   1118: 'Carrier 17 Power unit: Phase failure motor cable', class No Acknowledgement, trigger "DB302_HMI_Faults_Carrier17_Faults_1" bit 13
   1119: 'Carrier 17 Power unit: Ground fault', class No Acknowledgement, trigger "DB302_HMI_Faults_Carrier17_Faults_1" bit 14
   1120: 'Spare_Fault_1120', class No Acknowledgement, trigger "DB302_HMI_Faults_Carrier17_Faults_1" bit 15
   1121: 'Carrier 17 Motion Off Fault', class No Acknowledgement, trigger "DB302_HMI_Faults_Carrier17_Faults_2" bit 0
   1122: 'Carrier 17 Motion On Fault', class No Acknowledgement, trigger "DB302_HMI_Faults_Carrier17_Faults_2" bit 1
   1123: 'Carrier 17 Spacing Fault', class No Acknowledgement, trigger "DB302_HMI_Faults_Carrier17_Faults_2" bit 2
   1124: 'Carrier 17 Duplicate Carrier Number Fault', class No Acknowledgement, trigger "DB302_HMI_Faults_Carrier17_Faults_2" bit 3
   1125: 'Spare_Fault_1125', class No Acknowledgement, trigger "DB302_HMI_Faults_Carrier17_Faults_2" bit 4
   1126: 'Spare_Fault_1126', class No Acknowledgement, trigger "DB302_HMI_Faults_Carrier17_Faults_2" bit 5
   1127: 'Spare_Fault_1127', class No Acknowledgement, trigger "DB302_HMI_Faults_Carrier17_Faults_2" bit 6
   1128: 'Spare_Fault_1128', class No Acknowledgement, trigger "DB302_HMI_Faults_Carrier17_Faults_2" bit 7
   1129: 'Spare_Fault_1129', class No Acknowledgement, trigger "DB302_HMI_Faults_Carrier17_Faults_2" bit 8
   1130: 'Spare_Fault_1130', class No Acknowledgement, trigger "DB302_HMI_Faults_Carrier17_Faults_2" bit 9
   1131: 'Spare_Fault_1131', class No Acknowledgement, trigger "DB302_HMI_Faults_Carrier17_Faults_2" bit 10
   1132: 'Spare_Fault_1132', class No Acknowledgement, trigger "DB302_HMI_Faults_Carrier17_Faults_2" bit 11
   1133: 'Spare_Fault_1133', class No Acknowledgement, trigger "DB302_HMI_Faults_Carrier17_Faults_2" bit 12
   1134: 'Spare_Fault_1134', class No Acknowledgement, trigger "DB302_HMI_Faults_Carrier17_Faults_2" bit 13
   1135: 'Spare_Fault_1135', class No Acknowledgement, trigger "DB302_HMI_Faults_Carrier17_Faults_2" bit 14
   1136: 'Spare_Fault_1136', class No Acknowledgement, trigger "DB302_HMI_Faults_Carrier17_Faults_2" bit 15
   1137: 'Spare_Fault_1137', class No Acknowledgement, trigger "DB302_HMI_Faults_Carrier17_Faults_3" bit 0
   1138: 'Spare_Fault_1138', class No Acknowledgement, trigger "DB302_HMI_Faults_Carrier17_Faults_3" bit 1
   1139: 'Spare_Fault_1139', class No Acknowledgement, trigger "DB302_HMI_Faults_Carrier17_Faults_3" bit 2
   1140: 'Spare_Fault_1140', class No Acknowledgement, trigger "DB302_HMI_Faults_Carrier17_Faults_3" bit 3
   1141: 'Spare_Fault_1141', class No Acknowledgement, trigger "DB302_HMI_Faults_Carrier17_Faults_3" bit 4
   1142: 'Spare_Fault_1142', class No Acknowledgement, trigger "DB302_HMI_Faults_Carrier17_Faults_3" bit 5
   1143: 'Spare_Fault_1143', class No Acknowledgement, trigger "DB302_HMI_Faults_Carrier17_Faults_3" bit 6
   1144: 'Spare_Fault_1144', class No Acknowledgement, trigger "DB302_HMI_Faults_Carrier17_Faults_3" bit 7
   1145: 'Spare_Fault_1145', class No Acknowledgement, trigger "DB302_HMI_Faults_Carrier17_Faults_3" bit 8
   1146: 'Spare_Fault_1146', class No Acknowledgement, trigger "DB302_HMI_Faults_Carrier17_Faults_3" bit 9
   1147: 'Spare_Fault_1147', class No Acknowledgement, trigger "DB302_HMI_Faults_Carrier17_Faults_3" bit 10
   1148: 'Spare_Fault_1148', class No Acknowledgement, trigger "DB302_HMI_Faults_Carrier17_Faults_3" bit 11
   1149: 'Spare_Fault_1149', class No Acknowledgement, trigger "DB302_HMI_Faults_Carrier17_Faults_3" bit 12
   1150: 'Spare_Fault_1150', class No Acknowledgement, trigger "DB302_HMI_Faults_Carrier17_Faults_3" bit 13
   1151: 'Spare_Fault_1151', class No Acknowledgement, trigger "DB302_HMI_Faults_Carrier17_Faults_3" bit 14
   1152: 'Spare_Fault_1152', class No Acknowledgement, trigger "DB302_HMI_Faults_Carrier17_Faults_3" bit 15
   1153: 'Carrier 18 Disconnect Open Power Fault DI11.0', class No Acknowledgement, trigger "DB302_HMI_Faults_Carrier18_Faults_0" bit 0
   1154: 'Carrier 18 Drive Profinet Comm Fault', class No Acknowledgement, trigger "DB302_HMI_Faults_Carrier18_Faults_0" bit 1
   1155: 'Carrier 18 Production Stop Not Reset', class No Acknowledgement, trigger "DB302_HMI_Faults_Carrier18_Faults_0" bit 2
   1156: 'Carrier 18 CB02122 Tripped', class No Acknowledgement, trigger "DB302_HMI_Faults_Carrier18_Faults_0" bit 3
   1157: 'Carrier 18 CB02123 Tripped', class No Acknowledgement, trigger "DB302_HMI_Faults_Carrier18_Faults_0" bit 4
   1158: 'Carrier 18 AUX1 CB Tripped', class No Acknowledgement, trigger "DB302_HMI_Faults_Carrier18_Faults_0" bit 5
   1159: 'Carrier 18 AUX2 CB Tripped', class No Acknowledgement, trigger "DB302_HMI_Faults_Carrier18_Faults_0" bit 6
   1160: 'Carrier 18 PLC Not Communicating', class No Acknowledgement, trigger "DB302_HMI_Faults_Carrier18_Faults_0" bit 7
   1161: 'Carrier 18 Safe Input Card Fault', class No Acknowledgement, trigger "DB302_HMI_Faults_Carrier18_Faults_0" bit 8
   1162: 'Carrier 18 Safe Output Card Fault', class No Acknowledgement, trigger "DB302_HMI_Faults_Carrier18_Faults_0" bit 9
   1163: 'Carrier 18 Standard Input Card Fault', class No Acknowledgement, trigger "DB302_HMI_Faults_Carrier18_Faults_0" bit 10
   1164: 'Carrier 18 Standard Output Card Fault', class No Acknowledgement, trigger "DB302_HMI_Faults_Carrier18_Faults_0" bit 11
   1165: 'Carrier 18 Encoder Position Fault', class No Acknowledgement, trigger "DB302_HMI_Faults_Carrier18_Faults_0" bit 12
   1166: 'Carrier 18 Encoder Internal Error', class No Acknowledgement, trigger "DB302_HMI_Faults_Carrier18_Faults_0" bit 13
   1167: 'Carrier 18 Encoder Comm Fault', class No Acknowledgement, trigger "DB302_HMI_Faults_Carrier18_Faults_0" bit 14
   1168: 'Carrier 18 HMI Comm Fault', class No Acknowledgement, trigger "DB302_HMI_Faults_Carrier18_Faults_0" bit 15
   1169: 'Carrier 18 Crash Detection Fault', class No Acknowledgement, trigger "DB302_HMI_Faults_Carrier18_Faults_1" bit 0
   1170: 'Carrier 18 Carrier Number Invalid', class No Acknowledgement, trigger "DB302_HMI_Faults_Carrier18_Faults_1" bit 1
   1171: 'Carrier 18 Drive: PROFINET configuration error', class No Acknowledgement, trigger "DB302_HMI_Faults_Carrier18_Faults_1" bit 2
   1172: 'Carrier 18 Drive: Error internal communications', class No Acknowledgement, trigger "DB302_HMI_Faults_Carrier18_Faults_1" bit 3
   1173: 'Carrier 18 Drive: Motor overtemperature', class No Acknowledgement, trigger "DB302_HMI_Faults_Carrier18_Faults_1" bit 4
   1174: 'Carrier 18 Drive: Motor overcurrent', class No Acknowledgement, trigger "DB302_HMI_Faults_Carrier18_Faults_1" bit 5
   1175: 'Carrier 18 Drive: Infeed or power unit not ready', class No Acknowledgement, trigger "DB302_HMI_Faults_Carrier18_Faults_1" bit 6
   1176: 'Carrier 18 Drive: Short-circuit/ground fault detected', class No Acknowledgement, trigger "DB302_HMI_Faults_Carrier18_Faults_1" bit 7
   1177: 'Carrier 18 Drive: PROFINET Setpoint timeout', class No Acknowledgement, trigger "DB302_HMI_Faults_Carrier18_Faults_1" bit 8
   1178: 'Carrier 18 Power unit: Overcurrent', class No Acknowledgement, trigger "DB302_HMI_Faults_Carrier18_Faults_1" bit 9
   1179: 'Carrier 18 Power unit: DC link voltage overvoltage', class No Acknowledgement, trigger "DB302_HMI_Faults_Carrier18_Faults_1" bit 10
   1180: 'Carrier 18 Power unit: DC link voltage undervoltage', class No Acknowledgement, trigger "DB302_HMI_Faults_Carrier18_Faults_1" bit 11
   1181: 'Carrier 18 Power unit: Line phase failure in main circuit', class No Acknowledgement, trigger "DB302_HMI_Faults_Carrier18_Faults_1" bit 12
   1182: 'Carrier 18 Power unit: Phase failure motor cable', class No Acknowledgement, trigger "DB302_HMI_Faults_Carrier18_Faults_1" bit 13
   1183: 'Carrier 18 Power unit: Ground fault', class No Acknowledgement, trigger "DB302_HMI_Faults_Carrier18_Faults_1" bit 14
   1184: 'Spare_Fault_1184', class No Acknowledgement, trigger "DB302_HMI_Faults_Carrier18_Faults_1" bit 15
   1185: 'Carrier 18 Motion Off Fault', class No Acknowledgement, trigger "DB302_HMI_Faults_Carrier18_Faults_2" bit 0
   1186: 'Carrier 18 Motion On Fault', class No Acknowledgement, trigger "DB302_HMI_Faults_Carrier18_Faults_2" bit 1
   1187: 'Carrier 18 Spacing Fault', class No Acknowledgement, trigger "DB302_HMI_Faults_Carrier18_Faults_2" bit 2
   1188: 'Carrier 18 Duplicate Carrier Number Fault', class No Acknowledgement, trigger "DB302_HMI_Faults_Carrier18_Faults_2" bit 3
   1189: 'Spare_Fault_1189', class No Acknowledgement, trigger "DB302_HMI_Faults_Carrier18_Faults_2" bit 4
   1190: 'Spare_Fault_1190', class No Acknowledgement, trigger "DB302_HMI_Faults_Carrier18_Faults_2" bit 5
   1191: 'Spare_Fault_1191', class No Acknowledgement, trigger "DB302_HMI_Faults_Carrier18_Faults_2" bit 6
   1192: 'Spare_Fault_1192', class No Acknowledgement, trigger "DB302_HMI_Faults_Carrier18_Faults_2" bit 7
   1193: 'Spare_Fault_1193', class No Acknowledgement, trigger "DB302_HMI_Faults_Carrier18_Faults_2" bit 8
   1194: 'Spare_Fault_1194', class No Acknowledgement, trigger "DB302_HMI_Faults_Carrier18_Faults_2" bit 9
   1195: 'Spare_Fault_1195', class No Acknowledgement, trigger "DB302_HMI_Faults_Carrier18_Faults_2" bit 10
   1196: 'Spare_Fault_1196', class No Acknowledgement, trigger "DB302_HMI_Faults_Carrier18_Faults_2" bit 11
   1197: 'Spare_Fault_1197', class No Acknowledgement, trigger "DB302_HMI_Faults_Carrier18_Faults_2" bit 12
   1198: 'Spare_Fault_1198', class No Acknowledgement, trigger "DB302_HMI_Faults_Carrier18_Faults_2" bit 13
   1199: 'Spare_Fault_1199', class No Acknowledgement, trigger "DB302_HMI_Faults_Carrier18_Faults_2" bit 14
   1200: 'Spare_Fault_1200', class No Acknowledgement, trigger "DB302_HMI_Faults_Carrier18_Faults_2" bit 15
   1201: 'Spare_Fault_1201', class No Acknowledgement, trigger "DB302_HMI_Faults_Carrier18_Faults_3" bit 0
   1202: 'Spare_Fault_1202', class No Acknowledgement, trigger "DB302_HMI_Faults_Carrier18_Faults_3" bit 1
   1203: 'Spare_Fault_1203', class No Acknowledgement, trigger "DB302_HMI_Faults_Carrier18_Faults_3" bit 2
   1204: 'Spare_Fault_1204', class No Acknowledgement, trigger "DB302_HMI_Faults_Carrier18_Faults_3" bit 3
   1205: 'Spare_Fault_1205', class No Acknowledgement, trigger "DB302_HMI_Faults_Carrier18_Faults_3" bit 4
   1206: 'Spare_Fault_1206', class No Acknowledgement, trigger "DB302_HMI_Faults_Carrier18_Faults_3" bit 5
   1207: 'Spare_Fault_1207', class No Acknowledgement, trigger "DB302_HMI_Faults_Carrier18_Faults_3" bit 6
   1208: 'Spare_Fault_1208', class No Acknowledgement, trigger "DB302_HMI_Faults_Carrier18_Faults_3" bit 7
   1209: 'Spare_Fault_1209', class No Acknowledgement, trigger "DB302_HMI_Faults_Carrier18_Faults_3" bit 8
   1210: 'Spare_Fault_1210', class No Acknowledgement, trigger "DB302_HMI_Faults_Carrier18_Faults_3" bit 9
   1211: 'Spare_Fault_1211', class No Acknowledgement, trigger "DB302_HMI_Faults_Carrier18_Faults_3" bit 10
   1212: 'Spare_Fault_1212', class No Acknowledgement, trigger "DB302_HMI_Faults_Carrier18_Faults_3" bit 11
   1213: 'Spare_Fault_1213', class No Acknowledgement, trigger "DB302_HMI_Faults_Carrier18_Faults_3" bit 12
   1214: 'Spare_Fault_1214', class No Acknowledgement, trigger "DB302_HMI_Faults_Carrier18_Faults_3" bit 13
   1215: 'Spare_Fault_1215', class No Acknowledgement, trigger "DB302_HMI_Faults_Carrier18_Faults_3" bit 14
   1216: 'Spare_Fault_1216', class No Acknowledgement, trigger "DB302_HMI_Faults_Carrier18_Faults_3" bit 15
   1217: 'Carrier 19 Disconnect Open Power Fault DI11.0', class No Acknowledgement, trigger "DB302_HMI_Faults_Carrier19_Faults_0" bit 0
   1218: 'Carrier 19 Drive Profinet Comm Fault', class No Acknowledgement, trigger "DB302_HMI_Faults_Carrier19_Faults_0" bit 1
   1219: 'Carrier 19 Production Stop Not Reset', class No Acknowledgement, trigger "DB302_HMI_Faults_Carrier19_Faults_0" bit 2
   1220: 'Carrier 19 CB02122 Tripped', class No Acknowledgement, trigger "DB302_HMI_Faults_Carrier19_Faults_0" bit 3
   1221: 'Carrier 19 CB02123 Tripped', class No Acknowledgement, trigger "DB302_HMI_Faults_Carrier19_Faults_0" bit 4
   1222: 'Carrier 19 AUX1 CB Tripped', class No Acknowledgement, trigger "DB302_HMI_Faults_Carrier19_Faults_0" bit 5
   1223: 'Carrier 19 AUX2 CB Tripped', class No Acknowledgement, trigger "DB302_HMI_Faults_Carrier19_Faults_0" bit 6
   1224: 'Carrier 19 PLC Not Communicating', class No Acknowledgement, trigger "DB302_HMI_Faults_Carrier19_Faults_0" bit 7
   1225: 'Carrier 19 Safe Input Card Fault', class No Acknowledgement, trigger "DB302_HMI_Faults_Carrier19_Faults_0" bit 8
   1226: 'Carrier 19 Safe Output Card Fault', class No Acknowledgement, trigger "DB302_HMI_Faults_Carrier19_Faults_0" bit 9
   1227: 'Carrier 19 Standard Input Card Fault', class No Acknowledgement, trigger "DB302_HMI_Faults_Carrier19_Faults_0" bit 10
   1228: 'Carrier 19 Standard Output Card Fault', class No Acknowledgement, trigger "DB302_HMI_Faults_Carrier19_Faults_0" bit 11
   1229: 'Carrier 19 Encoder Position Fault', class No Acknowledgement, trigger "DB302_HMI_Faults_Carrier19_Faults_0" bit 12
   1230: 'Carrier 19 Encoder Internal Error', class No Acknowledgement, trigger "DB302_HMI_Faults_Carrier19_Faults_0" bit 13
   1231: 'Carrier 19 Encoder Comm Fault', class No Acknowledgement, trigger "DB302_HMI_Faults_Carrier19_Faults_0" bit 14
   1232: 'Carrier 19 HMI Comm Fault', class No Acknowledgement, trigger "DB302_HMI_Faults_Carrier19_Faults_0" bit 15
   1233: 'Carrier 19 Crash Detection Fault', class No Acknowledgement, trigger "DB302_HMI_Faults_Carrier19_Faults_1" bit 0
   1234: 'Carrier 19 Carrier Number Invalid', class No Acknowledgement, trigger "DB302_HMI_Faults_Carrier19_Faults_1" bit 1
   1235: 'Carrier 19 Drive: PROFINET configuration error', class No Acknowledgement, trigger "DB302_HMI_Faults_Carrier19_Faults_1" bit 2
   1236: 'Carrier 19 Drive: Error internal communications', class No Acknowledgement, trigger "DB302_HMI_Faults_Carrier19_Faults_1" bit 3
   1237: 'Carrier 19 Drive: Motor overtemperature', class No Acknowledgement, trigger "DB302_HMI_Faults_Carrier19_Faults_1" bit 4
   1238: 'Carrier 19 Drive: Motor overcurrent', class No Acknowledgement, trigger "DB302_HMI_Faults_Carrier19_Faults_1" bit 5
   1239: 'Carrier 19 Drive: Infeed or power unit not ready', class No Acknowledgement, trigger "DB302_HMI_Faults_Carrier19_Faults_1" bit 6
   1240: 'Carrier 19 Drive: Short-circuit/ground fault detected', class No Acknowledgement, trigger "DB302_HMI_Faults_Carrier19_Faults_1" bit 7
   1241: 'Carrier 19 Drive: PROFINET Setpoint timeout', class No Acknowledgement, trigger "DB302_HMI_Faults_Carrier19_Faults_1" bit 8
   1242: 'Carrier 19 Power unit: Overcurrent', class No Acknowledgement, trigger "DB302_HMI_Faults_Carrier19_Faults_1" bit 9
   1243: 'Carrier 19 Power unit: DC link voltage overvoltage', class No Acknowledgement, trigger "DB302_HMI_Faults_Carrier19_Faults_1" bit 10
   1244: 'Carrier 19 Power unit: DC link voltage undervoltage', class No Acknowledgement, trigger "DB302_HMI_Faults_Carrier19_Faults_1" bit 11
   1245: 'Carrier 19 Power unit: Line phase failure in main circuit', class No Acknowledgement, trigger "DB302_HMI_Faults_Carrier19_Faults_1" bit 12
   1246: 'Carrier 19 Power unit: Phase failure motor cable', class No Acknowledgement, trigger "DB302_HMI_Faults_Carrier19_Faults_1" bit 13
   1247: 'Carrier 19 Power unit: Ground fault', class No Acknowledgement, trigger "DB302_HMI_Faults_Carrier19_Faults_1" bit 14
   1248: 'Spare_Fault_1248', class No Acknowledgement, trigger "DB302_HMI_Faults_Carrier19_Faults_1" bit 15
   1249: 'Carrier 19 Motion Off Fault', class No Acknowledgement, trigger "DB302_HMI_Faults_Carrier19_Faults_2" bit 0
   1250: 'Carrier 19 Motion On Fault', class No Acknowledgement, trigger "DB302_HMI_Faults_Carrier19_Faults_2" bit 1
   1251: 'Carrier 19 Spacing Fault', class No Acknowledgement, trigger "DB302_HMI_Faults_Carrier19_Faults_2" bit 2
   1252: 'Carrier 19 Duplicate Carrier Number Fault', class No Acknowledgement, trigger "DB302_HMI_Faults_Carrier19_Faults_2" bit 3
   1253: 'Spare_Fault_1253', class No Acknowledgement, trigger "DB302_HMI_Faults_Carrier19_Faults_2" bit 4
   1254: 'Spare_Fault_1254', class No Acknowledgement, trigger "DB302_HMI_Faults_Carrier19_Faults_2" bit 5
   1255: 'Spare_Fault_1255', class No Acknowledgement, trigger "DB302_HMI_Faults_Carrier19_Faults_2" bit 6
   1256: 'Spare_Fault_1256', class No Acknowledgement, trigger "DB302_HMI_Faults_Carrier19_Faults_2" bit 7
   1257: 'Spare_Fault_1257', class No Acknowledgement, trigger "DB302_HMI_Faults_Carrier19_Faults_2" bit 8
   1258: 'Spare_Fault_1258', class No Acknowledgement, trigger "DB302_HMI_Faults_Carrier19_Faults_2" bit 9
   1259: 'Spare_Fault_1259', class No Acknowledgement, trigger "DB302_HMI_Faults_Carrier19_Faults_2" bit 10
   1260: 'Spare_Fault_1260', class No Acknowledgement, trigger "DB302_HMI_Faults_Carrier19_Faults_2" bit 11
   1261: 'Spare_Fault_1261', class No Acknowledgement, trigger "DB302_HMI_Faults_Carrier19_Faults_2" bit 12
   1262: 'Spare_Fault_1262', class No Acknowledgement, trigger "DB302_HMI_Faults_Carrier19_Faults_2" bit 13
   1263: 'Spare_Fault_1263', class No Acknowledgement, trigger "DB302_HMI_Faults_Carrier19_Faults_2" bit 14
   1264: 'Spare_Fault_1264', class No Acknowledgement, trigger "DB302_HMI_Faults_Carrier19_Faults_2" bit 15
   1265: 'Spare_Fault_1265', class No Acknowledgement, trigger "DB302_HMI_Faults_Carrier19_Faults_3" bit 0
   1266: 'Spare_Fault_1266', class No Acknowledgement, trigger "DB302_HMI_Faults_Carrier19_Faults_3" bit 1
   1267: 'Spare_Fault_1267', class No Acknowledgement, trigger "DB302_HMI_Faults_Carrier19_Faults_3" bit 2
   1268: 'Spare_Fault_1268', class No Acknowledgement, trigger "DB302_HMI_Faults_Carrier19_Faults_3" bit 3
   1269: 'Spare_Fault_1269', class No Acknowledgement, trigger "DB302_HMI_Faults_Carrier19_Faults_3" bit 4
   1270: 'Spare_Fault_1270', class No Acknowledgement, trigger "DB302_HMI_Faults_Carrier19_Faults_3" bit 5
   1271: 'Spare_Fault_1271', class No Acknowledgement, trigger "DB302_HMI_Faults_Carrier19_Faults_3" bit 6
   1272: 'Spare_Fault_1272', class No Acknowledgement, trigger "DB302_HMI_Faults_Carrier19_Faults_3" bit 7
   1273: 'Spare_Fault_1273', class No Acknowledgement, trigger "DB302_HMI_Faults_Carrier19_Faults_3" bit 8
   1274: 'Spare_Fault_1274', class No Acknowledgement, trigger "DB302_HMI_Faults_Carrier19_Faults_3" bit 9
   1275: 'Spare_Fault_1275', class No Acknowledgement, trigger "DB302_HMI_Faults_Carrier19_Faults_3" bit 10
   1276: 'Spare_Fault_1276', class No Acknowledgement, trigger "DB302_HMI_Faults_Carrier19_Faults_3" bit 11
   1277: 'Spare_Fault_1277', class No Acknowledgement, trigger "DB302_HMI_Faults_Carrier19_Faults_3" bit 12
   1278: 'Spare_Fault_1278', class No Acknowledgement, trigger "DB302_HMI_Faults_Carrier19_Faults_3" bit 13
   1279: 'Spare_Fault_1279', class No Acknowledgement, trigger "DB302_HMI_Faults_Carrier19_Faults_3" bit 14
   1280: 'Spare_Fault_1280', class No Acknowledgement, trigger "DB302_HMI_Faults_Carrier19_Faults_3" bit 15
   1281: 'Carrier 20 Disconnect Open Power Fault DI11.0', class No Acknowledgement, trigger "DB302_HMI_Faults_Carrier20_Faults_0" bit 0
   1282: 'Carrier 20 Drive Profinet Comm Fault', class No Acknowledgement, trigger "DB302_HMI_Faults_Carrier20_Faults_0" bit 1
   1283: 'Carrier 20 Production Stop Not Reset', class No Acknowledgement, trigger "DB302_HMI_Faults_Carrier20_Faults_0" bit 2
   1284: 'Carrier 20 CB02122 Tripped', class No Acknowledgement, trigger "DB302_HMI_Faults_Carrier20_Faults_0" bit 3
   1285: 'Carrier 20 CB02123 Tripped', class No Acknowledgement, trigger "DB302_HMI_Faults_Carrier20_Faults_0" bit 4
   1286: 'Carrier 20 AUX1 CB Tripped', class No Acknowledgement, trigger "DB302_HMI_Faults_Carrier20_Faults_0" bit 5
   1287: 'Carrier 20 AUX2 CB Tripped', class No Acknowledgement, trigger "DB302_HMI_Faults_Carrier20_Faults_0" bit 6
   1288: 'Carrier 20 PLC Not Communicating', class No Acknowledgement, trigger "DB302_HMI_Faults_Carrier20_Faults_0" bit 7
   1289: 'Carrier 20 Safe Input Card Fault', class No Acknowledgement, trigger "DB302_HMI_Faults_Carrier20_Faults_0" bit 8
   1290: 'Carrier 20 Safe Output Card Fault', class No Acknowledgement, trigger "DB302_HMI_Faults_Carrier20_Faults_0" bit 9
   1291: 'Carrier 20 Standard Input Card Fault', class No Acknowledgement, trigger "DB302_HMI_Faults_Carrier20_Faults_0" bit 10
   1292: 'Carrier 20 Standard Output Card Fault', class No Acknowledgement, trigger "DB302_HMI_Faults_Carrier20_Faults_0" bit 11
   1293: 'Carrier 20 Encoder Position Fault', class No Acknowledgement, trigger "DB302_HMI_Faults_Carrier20_Faults_0" bit 12
   1294: 'Carrier 20 Encoder Internal Error', class No Acknowledgement, trigger "DB302_HMI_Faults_Carrier20_Faults_0" bit 13
   1295: 'Carrier 20 Encoder Comm Fault', class No Acknowledgement, trigger "DB302_HMI_Faults_Carrier20_Faults_0" bit 14
   1296: 'Carrier 20 HMI Comm Fault', class No Acknowledgement, trigger "DB302_HMI_Faults_Carrier20_Faults_0" bit 15
   1297: 'Carrier 20 Crash Detection Fault', class No Acknowledgement, trigger "DB302_HMI_Faults_Carrier20_Faults_1" bit 0
   1298: 'Carrier 20 Carrier Number Invalid', class No Acknowledgement, trigger "DB302_HMI_Faults_Carrier20_Faults_1" bit 1
   1299: 'Carrier 20 Drive: PROFINET configuration error', class No Acknowledgement, trigger "DB302_HMI_Faults_Carrier20_Faults_1" bit 2
   1300: 'Carrier 20 Drive: Error internal communications', class No Acknowledgement, trigger "DB302_HMI_Faults_Carrier20_Faults_1" bit 3
   1301: 'Carrier 20 Drive: Motor overtemperature', class No Acknowledgement, trigger "DB302_HMI_Faults_Carrier20_Faults_1" bit 4
   1302: 'Carrier 20 Drive: Motor overcurrent', class No Acknowledgement, trigger "DB302_HMI_Faults_Carrier20_Faults_1" bit 5
   1303: 'Carrier 20 Drive: Infeed or power unit not ready', class No Acknowledgement, trigger "DB302_HMI_Faults_Carrier20_Faults_1" bit 6
   1304: 'Carrier 20 Drive: Short-circuit/ground fault detected', class No Acknowledgement, trigger "DB302_HMI_Faults_Carrier20_Faults_1" bit 7
   1305: 'Carrier 20 Drive: PROFINET Setpoint timeout', class No Acknowledgement, trigger "DB302_HMI_Faults_Carrier20_Faults_1" bit 8
   1306: 'Carrier 20 Power unit: Overcurrent', class No Acknowledgement, trigger "DB302_HMI_Faults_Carrier20_Faults_1" bit 9
   1307: 'Carrier 20 Power unit: DC link voltage overvoltage', class No Acknowledgement, trigger "DB302_HMI_Faults_Carrier20_Faults_1" bit 10
   1308: 'Carrier 20 Power unit: DC link voltage undervoltage', class No Acknowledgement, trigger "DB302_HMI_Faults_Carrier20_Faults_1" bit 11
   1309: 'Carrier 20 Power unit: Line phase failure in main circuit', class No Acknowledgement, trigger "DB302_HMI_Faults_Carrier20_Faults_1" bit 12
   1310: 'Carrier 20 Power unit: Phase failure motor cable', class No Acknowledgement, trigger "DB302_HMI_Faults_Carrier20_Faults_1" bit 13
   1311: 'Carrier 20 Power unit: Ground fault', class No Acknowledgement, trigger "DB302_HMI_Faults_Carrier20_Faults_1" bit 14
   1312: 'Spare_Fault_1312', class No Acknowledgement, trigger "DB302_HMI_Faults_Carrier20_Faults_1" bit 15
   1313: 'Carrier 20 Motion Off Fault', class No Acknowledgement, trigger "DB302_HMI_Faults_Carrier20_Faults_2" bit 0
   1314: 'Carrier 20 Motion On Fault', class No Acknowledgement, trigger "DB302_HMI_Faults_Carrier20_Faults_2" bit 1
   1315: 'Carrier 20 Spacing Fault', class No Acknowledgement, trigger "DB302_HMI_Faults_Carrier20_Faults_2" bit 2
   1316: 'Carrier 20 Duplicate Carrier Number Fault', class No Acknowledgement, trigger "DB302_HMI_Faults_Carrier20_Faults_2" bit 3
   1317: 'Spare_Fault_1317', class No Acknowledgement, trigger "DB302_HMI_Faults_Carrier20_Faults_2" bit 4
   1318: 'Spare_Fault_1318', class No Acknowledgement, trigger "DB302_HMI_Faults_Carrier20_Faults_2" bit 5
   1319: 'Spare_Fault_1319', class No Acknowledgement, trigger "DB302_HMI_Faults_Carrier20_Faults_2" bit 6
   1320: 'Spare_Fault_1320', class No Acknowledgement, trigger "DB302_HMI_Faults_Carrier20_Faults_2" bit 7
   1321: 'Spare_Fault_1321', class No Acknowledgement, trigger "DB302_HMI_Faults_Carrier20_Faults_2" bit 8
   1322: 'Spare_Fault_1322', class No Acknowledgement, trigger "DB302_HMI_Faults_Carrier20_Faults_2" bit 9
   1323: 'Spare_Fault_1323', class No Acknowledgement, trigger "DB302_HMI_Faults_Carrier20_Faults_2" bit 10
   1324: 'Spare_Fault_1324', class No Acknowledgement, trigger "DB302_HMI_Faults_Carrier20_Faults_2" bit 11
   1325: 'Spare_Fault_1325', class No Acknowledgement, trigger "DB302_HMI_Faults_Carrier20_Faults_2" bit 12
   1326: 'Spare_Fault_1326', class No Acknowledgement, trigger "DB302_HMI_Faults_Carrier20_Faults_2" bit 13
   1327: 'Spare_Fault_1327', class No Acknowledgement, trigger "DB302_HMI_Faults_Carrier20_Faults_2" bit 14
   1328: 'Spare_Fault_1328', class No Acknowledgement, trigger "DB302_HMI_Faults_Carrier20_Faults_2" bit 15
   1329: 'Spare_Fault_1329', class No Acknowledgement, trigger "DB302_HMI_Faults_Carrier20_Faults_3" bit 0
   1330: 'Spare_Fault_1330', class No Acknowledgement, trigger "DB302_HMI_Faults_Carrier20_Faults_3" bit 1
   1331: 'Spare_Fault_1331', class No Acknowledgement, trigger "DB302_HMI_Faults_Carrier20_Faults_3" bit 2
   1332: 'Spare_Fault_1332', class No Acknowledgement, trigger "DB302_HMI_Faults_Carrier20_Faults_3" bit 3
   1333: 'Spare_Fault_1333', class No Acknowledgement, trigger "DB302_HMI_Faults_Carrier20_Faults_3" bit 4
   1334: 'Spare_Fault_1334', class No Acknowledgement, trigger "DB302_HMI_Faults_Carrier20_Faults_3" bit 5
   1335: 'Spare_Fault_1335', class No Acknowledgement, trigger "DB302_HMI_Faults_Carrier20_Faults_3" bit 6
   1336: 'Spare_Fault_1336', class No Acknowledgement, trigger "DB302_HMI_Faults_Carrier20_Faults_3" bit 7
   1337: 'Spare_Fault_1337', class No Acknowledgement, trigger "DB302_HMI_Faults_Carrier20_Faults_3" bit 8
   1338: 'Spare_Fault_1338', class No Acknowledgement, trigger "DB302_HMI_Faults_Carrier20_Faults_3" bit 9
   1339: 'Spare_Fault_1339', class No Acknowledgement, trigger "DB302_HMI_Faults_Carrier20_Faults_3" bit 10
   1340: 'Spare_Fault_1340', class No Acknowledgement, trigger "DB302_HMI_Faults_Carrier20_Faults_3" bit 11
   1341: 'Spare_Fault_1341', class No Acknowledgement, trigger "DB302_HMI_Faults_Carrier20_Faults_3" bit 12
   1342: 'Spare_Fault_1342', class No Acknowledgement, trigger "DB302_HMI_Faults_Carrier20_Faults_3" bit 13
   1343: 'Spare_Fault_1343', class No Acknowledgement, trigger "DB302_HMI_Faults_Carrier20_Faults_3" bit 14
   1344: 'Spare_Fault_1344', class No Acknowledgement, trigger "DB302_HMI_Faults_Carrier20_Faults_3" bit 15
   1345: 'Carrier 21 Disconnect Open Power Fault DI11.0', class No Acknowledgement, trigger "DB302_HMI_Faults_Carrier21_Faults_0" bit 0
   1346: 'Carrier 21 Drive Profinet Comm Fault', class No Acknowledgement, trigger "DB302_HMI_Faults_Carrier21_Faults_0" bit 1
   1347: 'Carrier 21 Production Stop Not Reset', class No Acknowledgement, trigger "DB302_HMI_Faults_Carrier21_Faults_0" bit 2
   1348: 'Carrier 21 CB02122 Tripped', class No Acknowledgement, trigger "DB302_HMI_Faults_Carrier21_Faults_0" bit 3
   1349: 'Carrier 21 CB02123 Tripped', class No Acknowledgement, trigger "DB302_HMI_Faults_Carrier21_Faults_0" bit 4
   1350: 'Carrier 21 AUX1 CB Tripped', class No Acknowledgement, trigger "DB302_HMI_Faults_Carrier21_Faults_0" bit 5
   1351: 'Carrier 21 AUX2 CB Tripped', class No Acknowledgement, trigger "DB302_HMI_Faults_Carrier21_Faults_0" bit 6
   1352: 'Carrier 21 PLC Not Communicating', class No Acknowledgement, trigger "DB302_HMI_Faults_Carrier21_Faults_0" bit 7
   1353: 'Carrier 21 Safe Input Card Fault', class No Acknowledgement, trigger "DB302_HMI_Faults_Carrier21_Faults_0" bit 8
   1354: 'Carrier 21 Safe Output Card Fault', class No Acknowledgement, trigger "DB302_HMI_Faults_Carrier21_Faults_0" bit 9
   1355: 'Carrier 21 Standard Input Card Fault', class No Acknowledgement, trigger "DB302_HMI_Faults_Carrier21_Faults_0" bit 10
   1356: 'Carrier 21 Standard Output Card Fault', class No Acknowledgement, trigger "DB302_HMI_Faults_Carrier21_Faults_0" bit 11
   1357: 'Carrier 21 Encoder Position Fault', class No Acknowledgement, trigger "DB302_HMI_Faults_Carrier21_Faults_0" bit 12
   1358: 'Carrier 21 Encoder Internal Error', class No Acknowledgement, trigger "DB302_HMI_Faults_Carrier21_Faults_0" bit 13
   1359: 'Carrier 21 Encoder Comm Fault', class No Acknowledgement, trigger "DB302_HMI_Faults_Carrier21_Faults_0" bit 14
   1360: 'Carrier 21 HMI Comm Fault', class No Acknowledgement, trigger "DB302_HMI_Faults_Carrier21_Faults_0" bit 15
   1361: 'Carrier 21 Crash Detection Fault', class No Acknowledgement, trigger "DB302_HMI_Faults_Carrier21_Faults_1" bit 0
   1362: 'Carrier 21 Carrier Number Invalid', class No Acknowledgement, trigger "DB302_HMI_Faults_Carrier21_Faults_1" bit 1
   1363: 'Carrier 21 Drive: PROFINET configuration error', class No Acknowledgement, trigger "DB302_HMI_Faults_Carrier21_Faults_1" bit 2
   1364: 'Carrier 21 Drive: Error internal communications', class No Acknowledgement, trigger "DB302_HMI_Faults_Carrier21_Faults_1" bit 3
   1365: 'Carrier 21 Drive: Motor overtemperature', class No Acknowledgement, trigger "DB302_HMI_Faults_Carrier21_Faults_1" bit 4
   1366: 'Carrier 21 Drive: Motor overcurrent', class No Acknowledgement, trigger "DB302_HMI_Faults_Carrier21_Faults_1" bit 5
   1367: 'Carrier 21 Drive: Infeed or power unit not ready', class No Acknowledgement, trigger "DB302_HMI_Faults_Carrier21_Faults_1" bit 6
   1368: 'Carrier 21 Drive: Short-circuit/ground fault detected', class No Acknowledgement, trigger "DB302_HMI_Faults_Carrier21_Faults_1" bit 7
   1369: 'Carrier 21 Drive: PROFINET Setpoint timeout', class No Acknowledgement, trigger "DB302_HMI_Faults_Carrier21_Faults_1" bit 8
   1370: 'Carrier 21 Power unit: Overcurrent', class No Acknowledgement, trigger "DB302_HMI_Faults_Carrier21_Faults_1" bit 9
   1371: 'Carrier 21 Power unit: DC link voltage overvoltage', class No Acknowledgement, trigger "DB302_HMI_Faults_Carrier21_Faults_1" bit 10
   1372: 'Carrier 21 Power unit: DC link voltage undervoltage', class No Acknowledgement, trigger "DB302_HMI_Faults_Carrier21_Faults_1" bit 11
   1373: 'Carrier 21 Power unit: Line phase failure in main circuit', class No Acknowledgement, trigger "DB302_HMI_Faults_Carrier21_Faults_1" bit 12
   1374: 'Carrier 21 Power unit: Phase failure motor cable', class No Acknowledgement, trigger "DB302_HMI_Faults_Carrier21_Faults_1" bit 13
   1375: 'Carrier 21 Power unit: Ground fault', class No Acknowledgement, trigger "DB302_HMI_Faults_Carrier21_Faults_1" bit 14
   1376: 'Spare_Fault_1376', class No Acknowledgement, trigger "DB302_HMI_Faults_Carrier21_Faults_1" bit 15
   1377: 'Carrier 21 Motion Off Fault', class No Acknowledgement, trigger "DB302_HMI_Faults_Carrier21_Faults_2" bit 0
   1378: 'Carrier 21 Motion On Fault', class No Acknowledgement, trigger "DB302_HMI_Faults_Carrier21_Faults_2" bit 1
   1379: 'Carrier 21 Spacing Fault', class No Acknowledgement, trigger "DB302_HMI_Faults_Carrier21_Faults_2" bit 2
   1380: 'Carrier 21 Duplicate Carrier Number Fault', class No Acknowledgement, trigger "DB302_HMI_Faults_Carrier21_Faults_2" bit 3
   1381: 'Spare_Fault_1381', class No Acknowledgement, trigger "DB302_HMI_Faults_Carrier21_Faults_2" bit 4
   1382: 'Spare_Fault_1382', class No Acknowledgement, trigger "DB302_HMI_Faults_Carrier21_Faults_2" bit 5
   1383: 'Spare_Fault_1383', class No Acknowledgement, trigger "DB302_HMI_Faults_Carrier21_Faults_2" bit 6
   1384: 'Spare_Fault_1384', class No Acknowledgement, trigger "DB302_HMI_Faults_Carrier21_Faults_2" bit 7
   1385: 'Spare_Fault_1385', class No Acknowledgement, trigger "DB302_HMI_Faults_Carrier21_Faults_2" bit 8
   1386: 'Spare_Fault_1386', class No Acknowledgement, trigger "DB302_HMI_Faults_Carrier21_Faults_2" bit 9
   1387: 'Spare_Fault_1387', class No Acknowledgement, trigger "DB302_HMI_Faults_Carrier21_Faults_2" bit 10
   1388: 'Spare_Fault_1388', class No Acknowledgement, trigger "DB302_HMI_Faults_Carrier21_Faults_2" bit 11
   1389: 'Spare_Fault_1389', class No Acknowledgement, trigger "DB302_HMI_Faults_Carrier21_Faults_2" bit 12
   1390: 'Spare_Fault_1390', class No Acknowledgement, trigger "DB302_HMI_Faults_Carrier21_Faults_2" bit 13
   1391: 'Spare_Fault_1391', class No Acknowledgement, trigger "DB302_HMI_Faults_Carrier21_Faults_2" bit 14
   1392: 'Spare_Fault_1392', class No Acknowledgement, trigger "DB302_HMI_Faults_Carrier21_Faults_2" bit 15
   1393: 'Spare_Fault_1393', class No Acknowledgement, trigger "DB302_HMI_Faults_Carrier21_Faults_3" bit 0
   1394: 'Spare_Fault_1394', class No Acknowledgement, trigger "DB302_HMI_Faults_Carrier21_Faults_3" bit 1
   1395: 'Spare_Fault_1395', class No Acknowledgement, trigger "DB302_HMI_Faults_Carrier21_Faults_3" bit 2
   1396: 'Spare_Fault_1396', class No Acknowledgement, trigger "DB302_HMI_Faults_Carrier21_Faults_3" bit 3
   1397: 'Spare_Fault_1397', class No Acknowledgement, trigger "DB302_HMI_Faults_Carrier21_Faults_3" bit 4
   1398: 'Spare_Fault_1398', class No Acknowledgement, trigger "DB302_HMI_Faults_Carrier21_Faults_3" bit 5
   1399: 'Spare_Fault_1399', class No Acknowledgement, trigger "DB302_HMI_Faults_Carrier21_Faults_3" bit 6
   1400: 'Spare_Fault_1400', class No Acknowledgement, trigger "DB302_HMI_Faults_Carrier21_Faults_3" bit 7
   1401: 'Spare_Fault_1401', class No Acknowledgement, trigger "DB302_HMI_Faults_Carrier21_Faults_3" bit 8
   1402: 'Spare_Fault_1402', class No Acknowledgement, trigger "DB302_HMI_Faults_Carrier21_Faults_3" bit 9
   1403: 'Spare_Fault_1403', class No Acknowledgement, trigger "DB302_HMI_Faults_Carrier21_Faults_3" bit 10
   1404: 'Spare_Fault_1404', class No Acknowledgement, trigger "DB302_HMI_Faults_Carrier21_Faults_3" bit 11
   1405: 'Spare_Fault_1405', class No Acknowledgement, trigger "DB302_HMI_Faults_Carrier21_Faults_3" bit 12
   1406: 'Spare_Fault_1406', class No Acknowledgement, trigger "DB302_HMI_Faults_Carrier21_Faults_3" bit 13
   1407: 'Spare_Fault_1407', class No Acknowledgement, trigger "DB302_HMI_Faults_Carrier21_Faults_3" bit 14
   1408: 'Spare_Fault_1408', class No Acknowledgement, trigger "DB302_HMI_Faults_Carrier21_Faults_3" bit 15
   1409: 'Carrier 22 Disconnect Open Power Fault DI11.0', class No Acknowledgement, trigger "DB302_HMI_Faults_Carrier22_Faults_0" bit 0
   1410: 'Carrier 22 Drive Profinet Comm Fault', class No Acknowledgement, trigger "DB302_HMI_Faults_Carrier22_Faults_0" bit 1
   1411: 'Carrier 22 Production Stop Not Reset', class No Acknowledgement, trigger "DB302_HMI_Faults_Carrier22_Faults_0" bit 2
   1412: 'Carrier 22 CB02122 Tripped', class No Acknowledgement, trigger "DB302_HMI_Faults_Carrier22_Faults_0" bit 3
   1413: 'Carrier 22 CB02123 Tripped', class No Acknowledgement, trigger "DB302_HMI_Faults_Carrier22_Faults_0" bit 4
   1414: 'Carrier 22 AUX1 CB Tripped', class No Acknowledgement, trigger "DB302_HMI_Faults_Carrier22_Faults_0" bit 5
   1415: 'Carrier 22 AUX2 CB Tripped', class No Acknowledgement, trigger "DB302_HMI_Faults_Carrier22_Faults_0" bit 6
   1416: 'Carrier 22 PLC Not Communicating', class No Acknowledgement, trigger "DB302_HMI_Faults_Carrier22_Faults_0" bit 7
   1417: 'Carrier 22 Safe Input Card Fault', class No Acknowledgement, trigger "DB302_HMI_Faults_Carrier22_Faults_0" bit 8
   1418: 'Carrier 22 Safe Output Card Fault', class No Acknowledgement, trigger "DB302_HMI_Faults_Carrier22_Faults_0" bit 9
   1419: 'Carrier 22 Standard Input Card Fault', class No Acknowledgement, trigger "DB302_HMI_Faults_Carrier22_Faults_0" bit 10
   1420: 'Carrier 22 Standard Output Card Fault', class No Acknowledgement, trigger "DB302_HMI_Faults_Carrier22_Faults_0" bit 11
   1421: 'Carrier 22 Encoder Position Fault', class No Acknowledgement, trigger "DB302_HMI_Faults_Carrier22_Faults_0" bit 12
   1422: 'Carrier 22 Encoder Internal Error', class No Acknowledgement, trigger "DB302_HMI_Faults_Carrier22_Faults_0" bit 13
   1423: 'Carrier 22 Encoder Comm Fault', class No Acknowledgement, trigger "DB302_HMI_Faults_Carrier22_Faults_0" bit 14
   1424: 'Carrier 22 HMI Comm Fault', class No Acknowledgement, trigger "DB302_HMI_Faults_Carrier22_Faults_0" bit 15
   1425: 'Carrier 22 Crash Detection Fault', class No Acknowledgement, trigger "DB302_HMI_Faults_Carrier22_Faults_1" bit 0
   1426: 'Carrier 22 Carrier Number Invalid', class No Acknowledgement, trigger "DB302_HMI_Faults_Carrier22_Faults_1" bit 1
   1427: 'Carrier 22 Drive: PROFINET configuration error', class No Acknowledgement, trigger "DB302_HMI_Faults_Carrier22_Faults_1" bit 2
   1428: 'Carrier 22 Drive: Error internal communications', class No Acknowledgement, trigger "DB302_HMI_Faults_Carrier22_Faults_1" bit 3
   1429: 'Carrier 22 Drive: Motor overtemperature', class No Acknowledgement, trigger "DB302_HMI_Faults_Carrier22_Faults_1" bit 4
   1430: 'Carrier 22 Drive: Motor overcurrent', class No Acknowledgement, trigger "DB302_HMI_Faults_Carrier22_Faults_1" bit 5
   1431: 'Carrier 22 Drive: Infeed or power unit not ready', class No Acknowledgement, trigger "DB302_HMI_Faults_Carrier22_Faults_1" bit 6
   1432: 'Carrier 22 Drive: Short-circuit/ground fault detected', class No Acknowledgement, trigger "DB302_HMI_Faults_Carrier22_Faults_1" bit 7
   1433: 'Carrier 22 Drive: PROFINET Setpoint timeout', class No Acknowledgement, trigger "DB302_HMI_Faults_Carrier22_Faults_1" bit 8
   1434: 'Carrier 22 Power unit: Overcurrent', class No Acknowledgement, trigger "DB302_HMI_Faults_Carrier22_Faults_1" bit 9
   1435: 'Carrier 22 Power unit: DC link voltage overvoltage', class No Acknowledgement, trigger "DB302_HMI_Faults_Carrier22_Faults_1" bit 10
   1436: 'Carrier 22 Power unit: DC link voltage undervoltage', class No Acknowledgement, trigger "DB302_HMI_Faults_Carrier22_Faults_1" bit 11
   1437: 'Carrier 22 Power unit: Line phase failure in main circuit', class No Acknowledgement, trigger "DB302_HMI_Faults_Carrier22_Faults_1" bit 12
   1438: 'Carrier 22 Power unit: Phase failure motor cable', class No Acknowledgement, trigger "DB302_HMI_Faults_Carrier22_Faults_1" bit 13
   1439: 'Carrier 22 Power unit: Ground fault', class No Acknowledgement, trigger "DB302_HMI_Faults_Carrier22_Faults_1" bit 14
   1440: 'Spare_Fault_1440', class No Acknowledgement, trigger "DB302_HMI_Faults_Carrier22_Faults_1" bit 15
   1441: 'Carrier 22 Motion Off Fault', class No Acknowledgement, trigger "DB302_HMI_Faults_Carrier22_Faults_2" bit 0
   1442: 'Carrier 22 Motion On Fault', class No Acknowledgement, trigger "DB302_HMI_Faults_Carrier22_Faults_2" bit 1
   1443: 'Carrier 22 Spacing Fault', class No Acknowledgement, trigger "DB302_HMI_Faults_Carrier22_Faults_2" bit 2
   1444: 'Carrier 22 Duplicate Carrier Number Fault', class No Acknowledgement, trigger "DB302_HMI_Faults_Carrier22_Faults_2" bit 3
   1445: 'Spare_Fault_1445', class No Acknowledgement, trigger "DB302_HMI_Faults_Carrier22_Faults_2" bit 4
   1446: 'Spare_Fault_1446', class No Acknowledgement, trigger "DB302_HMI_Faults_Carrier22_Faults_2" bit 5
   1447: 'Spare_Fault_1447', class No Acknowledgement, trigger "DB302_HMI_Faults_Carrier22_Faults_2" bit 6
   1448: 'Spare_Fault_1448', class No Acknowledgement, trigger "DB302_HMI_Faults_Carrier22_Faults_2" bit 7
   1449: 'Spare_Fault_1449', class No Acknowledgement, trigger "DB302_HMI_Faults_Carrier22_Faults_2" bit 8
   1450: 'Spare_Fault_1450', class No Acknowledgement, trigger "DB302_HMI_Faults_Carrier22_Faults_2" bit 9
   1451: 'Spare_Fault_1451', class No Acknowledgement, trigger "DB302_HMI_Faults_Carrier22_Faults_2" bit 10
   1452: 'Spare_Fault_1452', class No Acknowledgement, trigger "DB302_HMI_Faults_Carrier22_Faults_2" bit 11
   1453: 'Spare_Fault_1453', class No Acknowledgement, trigger "DB302_HMI_Faults_Carrier22_Faults_2" bit 12
   1454: 'Spare_Fault_1454', class No Acknowledgement, trigger "DB302_HMI_Faults_Carrier22_Faults_2" bit 13
   1455: 'Spare_Fault_1455', class No Acknowledgement, trigger "DB302_HMI_Faults_Carrier22_Faults_2" bit 14
   1456: 'Spare_Fault_1456', class No Acknowledgement, trigger "DB302_HMI_Faults_Carrier22_Faults_2" bit 15
   1457: 'Spare_Fault_1457', class No Acknowledgement, trigger "DB302_HMI_Faults_Carrier22_Faults_3" bit 0
   1458: 'Spare_Fault_1458', class No Acknowledgement, trigger "DB302_HMI_Faults_Carrier22_Faults_3" bit 1
   1459: 'Spare_Fault_1459', class No Acknowledgement, trigger "DB302_HMI_Faults_Carrier22_Faults_3" bit 2
   1460: 'Spare_Fault_1460', class No Acknowledgement, trigger "DB302_HMI_Faults_Carrier22_Faults_3" bit 3
   1461: 'Spare_Fault_1461', class No Acknowledgement, trigger "DB302_HMI_Faults_Carrier22_Faults_3" bit 4
   1462: 'Spare_Fault_1462', class No Acknowledgement, trigger "DB302_HMI_Faults_Carrier22_Faults_3" bit 5
   1463: 'Spare_Fault_1463', class No Acknowledgement, trigger "DB302_HMI_Faults_Carrier22_Faults_3" bit 6
   1464: 'Spare_Fault_1464', class No Acknowledgement, trigger "DB302_HMI_Faults_Carrier22_Faults_3" bit 7
   1465: 'Spare_Fault_1465', class No Acknowledgement, trigger "DB302_HMI_Faults_Carrier22_Faults_3" bit 8
   1466: 'Spare_Fault_1466', class No Acknowledgement, trigger "DB302_HMI_Faults_Carrier22_Faults_3" bit 9
   1467: 'Spare_Fault_1467', class No Acknowledgement, trigger "DB302_HMI_Faults_Carrier22_Faults_3" bit 10
   1468: 'Spare_Fault_1468', class No Acknowledgement, trigger "DB302_HMI_Faults_Carrier22_Faults_3" bit 11
   1469: 'Spare_Fault_1469', class No Acknowledgement, trigger "DB302_HMI_Faults_Carrier22_Faults_3" bit 12
   1470: 'Spare_Fault_1470', class No Acknowledgement, trigger "DB302_HMI_Faults_Carrier22_Faults_3" bit 13
   1471: 'Spare_Fault_1471', class No Acknowledgement, trigger "DB302_HMI_Faults_Carrier22_Faults_3" bit 14
   1472: 'Spare_Fault_1472', class No Acknowledgement, trigger "DB302_HMI_Faults_Carrier22_Faults_3" bit 15
   1473: 'Carrier 23 Disconnect Open Power Fault DI11.0', class No Acknowledgement, trigger "DB302_HMI_Faults_Carrier23_Faults_0" bit 0
   1474: 'Carrier 23 Drive Profinet Comm Fault', class No Acknowledgement, trigger "DB302_HMI_Faults_Carrier23_Faults_0" bit 1
   1475: 'Carrier 23 Production Stop Not Reset', class No Acknowledgement, trigger "DB302_HMI_Faults_Carrier23_Faults_0" bit 2
   1476: 'Carrier 23 CB02122 Tripped', class No Acknowledgement, trigger "DB302_HMI_Faults_Carrier23_Faults_0" bit 3
   1477: 'Carrier 23 CB02123 Tripped', class No Acknowledgement, trigger "DB302_HMI_Faults_Carrier23_Faults_0" bit 4
   1478: 'Carrier 23 AUX1 CB Tripped', class No Acknowledgement, trigger "DB302_HMI_Faults_Carrier23_Faults_0" bit 5
   1479: 'Carrier 23 AUX2 CB Tripped', class No Acknowledgement, trigger "DB302_HMI_Faults_Carrier23_Faults_0" bit 6
   1480: 'Carrier 23 PLC Not Communicating', class No Acknowledgement, trigger "DB302_HMI_Faults_Carrier23_Faults_0" bit 7
   1481: 'Carrier 23 Safe Input Card Fault', class No Acknowledgement, trigger "DB302_HMI_Faults_Carrier23_Faults_0" bit 8
   1482: 'Carrier 23 Safe Output Card Fault', class No Acknowledgement, trigger "DB302_HMI_Faults_Carrier23_Faults_0" bit 9
   1483: 'Carrier 23 Standard Input Card Fault', class No Acknowledgement, trigger "DB302_HMI_Faults_Carrier23_Faults_0" bit 10
   1484: 'Carrier 23 Standard Output Card Fault', class No Acknowledgement, trigger "DB302_HMI_Faults_Carrier23_Faults_0" bit 11
   1485: 'Carrier 23 Encoder Position Fault', class No Acknowledgement, trigger "DB302_HMI_Faults_Carrier23_Faults_0" bit 12
   1486: 'Carrier 23 Encoder Internal Error', class No Acknowledgement, trigger "DB302_HMI_Faults_Carrier23_Faults_0" bit 13
   1487: 'Carrier 23 Encoder Comm Fault', class No Acknowledgement, trigger "DB302_HMI_Faults_Carrier23_Faults_0" bit 14
   1488: 'Carrier 23 HMI Comm Fault', class No Acknowledgement, trigger "DB302_HMI_Faults_Carrier23_Faults_0" bit 15
   1489: 'Carrier 23 Crash Detection Fault', class No Acknowledgement, trigger "DB302_HMI_Faults_Carrier23_Faults_1" bit 0
   1490: 'Carrier 23 Carrier Number Invalid', class No Acknowledgement, trigger "DB302_HMI_Faults_Carrier23_Faults_1" bit 1
   1491: 'Carrier 23 Drive: PROFINET configuration error', class No Acknowledgement, trigger "DB302_HMI_Faults_Carrier23_Faults_1" bit 2
   1492: 'Carrier 23 Drive: Error internal communications', class No Acknowledgement, trigger "DB302_HMI_Faults_Carrier23_Faults_1" bit 3
   1493: 'Carrier 23 Drive: Motor overtemperature', class No Acknowledgement, trigger "DB302_HMI_Faults_Carrier23_Faults_1" bit 4
   1494: 'Carrier 23 Drive: Motor overcurrent', class No Acknowledgement, trigger "DB302_HMI_Faults_Carrier23_Faults_1" bit 5
   1495: 'Carrier 23 Drive: Infeed or power unit not ready', class No Acknowledgement, trigger "DB302_HMI_Faults_Carrier23_Faults_1" bit 6
   1496: 'Carrier 23 Drive: Short-circuit/ground fault detected', class No Acknowledgement, trigger "DB302_HMI_Faults_Carrier23_Faults_1" bit 7
   1497: 'Carrier 23 Drive: PROFINET Setpoint timeout', class No Acknowledgement, trigger "DB302_HMI_Faults_Carrier23_Faults_1" bit 8
   1498: 'Carrier 23 Power unit: Overcurrent', class No Acknowledgement, trigger "DB302_HMI_Faults_Carrier23_Faults_1" bit 9
   1499: 'Carrier 23 Power unit: DC link voltage overvoltage', class No Acknowledgement, trigger "DB302_HMI_Faults_Carrier23_Faults_1" bit 10
   1500: 'Carrier 23 Power unit: DC link voltage undervoltage', class No Acknowledgement, trigger "DB302_HMI_Faults_Carrier23_Faults_1" bit 11
   1501: 'Carrier 23 Power unit: Line phase failure in main circuit', class No Acknowledgement, trigger "DB302_HMI_Faults_Carrier23_Faults_1" bit 12
   1502: 'Carrier 23 Power unit: Phase failure motor cable', class No Acknowledgement, trigger "DB302_HMI_Faults_Carrier23_Faults_1" bit 13
   1503: 'Carrier 23 Power unit: Ground fault', class No Acknowledgement, trigger "DB302_HMI_Faults_Carrier23_Faults_1" bit 14
   1504: 'Spare_Fault_1504', class No Acknowledgement, trigger "DB302_HMI_Faults_Carrier23_Faults_1" bit 15
   1505: 'Carrier 23 Motion Off Fault', class No Acknowledgement, trigger "DB302_HMI_Faults_Carrier23_Faults_2" bit 0
   1506: 'Carrier 23 Motion On Fault', class No Acknowledgement, trigger "DB302_HMI_Faults_Carrier23_Faults_2" bit 1
   1507: 'Carrier 23 Spacing Fault', class No Acknowledgement, trigger "DB302_HMI_Faults_Carrier23_Faults_2" bit 2
   1508: 'Carrier 23 Duplicate Carrier Number Fault', class No Acknowledgement, trigger "DB302_HMI_Faults_Carrier23_Faults_2" bit 3
   1509: 'Spare_Fault_1509', class No Acknowledgement, trigger "DB302_HMI_Faults_Carrier23_Faults_2" bit 4
   1510: 'Spare_Fault_1510', class No Acknowledgement, trigger "DB302_HMI_Faults_Carrier23_Faults_2" bit 5
   1511: 'Spare_Fault_1511', class No Acknowledgement, trigger "DB302_HMI_Faults_Carrier23_Faults_2" bit 6
   1512: 'Spare_Fault_1512', class No Acknowledgement, trigger "DB302_HMI_Faults_Carrier23_Faults_2" bit 7
   1513: 'Spare_Fault_1513', class No Acknowledgement, trigger "DB302_HMI_Faults_Carrier23_Faults_2" bit 8
   1514: 'Spare_Fault_1514', class No Acknowledgement, trigger "DB302_HMI_Faults_Carrier23_Faults_2" bit 9
   1515: 'Spare_Fault_1515', class No Acknowledgement, trigger "DB302_HMI_Faults_Carrier23_Faults_2" bit 10
   1516: 'Spare_Fault_1516', class No Acknowledgement, trigger "DB302_HMI_Faults_Carrier23_Faults_2" bit 11
   1517: 'Spare_Fault_1517', class No Acknowledgement, trigger "DB302_HMI_Faults_Carrier23_Faults_2" bit 12
   1518: 'Spare_Fault_1518', class No Acknowledgement, trigger "DB302_HMI_Faults_Carrier23_Faults_2" bit 13
   1519: 'Spare_Fault_1519', class No Acknowledgement, trigger "DB302_HMI_Faults_Carrier23_Faults_2" bit 14
   1520: 'Spare_Fault_1520', class No Acknowledgement, trigger "DB302_HMI_Faults_Carrier23_Faults_2" bit 15
   1521: 'Spare_Fault_1521', class No Acknowledgement, trigger "DB302_HMI_Faults_Carrier23_Faults_3" bit 0
   1522: 'Spare_Fault_1522', class No Acknowledgement, trigger "DB302_HMI_Faults_Carrier23_Faults_3" bit 1
   1523: 'Spare_Fault_1523', class No Acknowledgement, trigger "DB302_HMI_Faults_Carrier23_Faults_3" bit 2
   1524: 'Spare_Fault_1524', class No Acknowledgement, trigger "DB302_HMI_Faults_Carrier23_Faults_3" bit 3
   1525: 'Spare_Fault_1525', class No Acknowledgement, trigger "DB302_HMI_Faults_Carrier23_Faults_3" bit 4
   1526: 'Spare_Fault_1526', class No Acknowledgement, trigger "DB302_HMI_Faults_Carrier23_Faults_3" bit 5
   1527: 'Spare_Fault_1527', class No Acknowledgement, trigger "DB302_HMI_Faults_Carrier23_Faults_3" bit 6
   1528: 'Spare_Fault_1528', class No Acknowledgement, trigger "DB302_HMI_Faults_Carrier23_Faults_3" bit 7
   1529: 'Spare_Fault_1529', class No Acknowledgement, trigger "DB302_HMI_Faults_Carrier23_Faults_3" bit 8
   1530: 'Spare_Fault_1530', class No Acknowledgement, trigger "DB302_HMI_Faults_Carrier23_Faults_3" bit 9
   1531: 'Spare_Fault_1531', class No Acknowledgement, trigger "DB302_HMI_Faults_Carrier23_Faults_3" bit 10
   1532: 'Spare_Fault_1532', class No Acknowledgement, trigger "DB302_HMI_Faults_Carrier23_Faults_3" bit 11
   1533: 'Spare_Fault_1533', class No Acknowledgement, trigger "DB302_HMI_Faults_Carrier23_Faults_3" bit 12
   1534: 'Spare_Fault_1534', class No Acknowledgement, trigger "DB302_HMI_Faults_Carrier23_Faults_3" bit 13
   1535: 'Spare_Fault_1535', class No Acknowledgement, trigger "DB302_HMI_Faults_Carrier23_Faults_3" bit 14
   1536: 'Spare_Fault_1536', class No Acknowledgement, trigger "DB302_HMI_Faults_Carrier23_Faults_3" bit 15
   1537: 'Carrier 24 Disconnect Open Power Fault DI11.0', class No Acknowledgement, trigger "DB302_HMI_Faults_Carrier24_Faults_0" bit 0
   1538: 'Carrier 24 Drive Profinet Comm Fault', class No Acknowledgement, trigger "DB302_HMI_Faults_Carrier24_Faults_0" bit 1
   1539: 'Carrier 24 Production Stop Not Reset', class No Acknowledgement, trigger "DB302_HMI_Faults_Carrier24_Faults_0" bit 2
   1540: 'Carrier 24 CB02122 Tripped', class No Acknowledgement, trigger "DB302_HMI_Faults_Carrier24_Faults_0" bit 3
